
     #error := false;
     #status := #STATUS_FINISHED_NO_ERROR;
     #subfunctionStatus := #SUB_STATUS_NO_ERROR;
     // ENO mechanism is not used
     ENO := TRUE;
   END_REGION
END_FUNCTION

FUNCTION "LGF_RandomRange_Real" : Real   // FC10014, SCL
TITLE = LGF_RandomRange_Real
{ S7_Optimized_Access := 'TRUE' }
AUTHOR : Siemens_Digital_Industries
FAMILY : LGF
NAME : LGF_RandomRange_Real
// This function generates random numbers in defined limits (Datatype Real)
   VAR_INPUT
      minValue : Real;   // minimal Value random can reach / Minimum value of the range of the random number
      maxValue : Real;   // maximal Value random can reach / Maximum value of the range of the random number
   END_VAR
   VAR_OUTPUT
      error : Bool;   // Error if true
      status : Word;   // Status of the function
      subfunctionStatus : Word;   // Status or return value of called FB's, FCs and system blocks
   END_VAR
   VAR_TEMP
      tempTime : DTL;   // System time
      tempNanoSecondInDWord : DWord;   // UDINT converted to DWORD for access to individual bytes
      tempTimeStatus : Word;   // Status of the instruction RD_SYS_T
      tempRandomValue : DWord;   // Random-start-value
      tempNormReal : Real;   // normalized value
   END_VAR
   // Ret_Val : Returns random Real number in predefined range
   VAR CONSTANT
      ZERO : Real := 0.0;   // Zero value in case of error
      MAX_UDINT : UDInt := 4294967295;   // Maximum UDINT value
      SUB_STATUS_NO_ERROR : Word := 16#0000;   // Status: sub function call ends without error
      STATUS_FINISHED_NO_ERROR : Word := 16#0000;   // Status: Execution finished without errors
      ERR_MAX_LESS_MIN : Word := 16#8200;   // Error: The maximum limit number is smaller than the minimum limit number
      ERR_RD_SYS_T : Word := 16#8600;   // Error: System function Read system time returned an error
   END_VAR
BEGIN
   REGION Block info header
     //=============================================================================
     // SIEMENS AG / (c)Copyright 2017
     //-----------------------------------------------------------------------------
     // Title:            LGF_RandomRange_Real
     // Comment/Function: This function generates random numbers in defined limits (Datatype Real)
     // Library/Family:   LGF(Library General Functions)
     // Author:           Siemens Digital Industry Support
     // Tested with:      S7-PLCSIM Advanced V2.0 SP1
     // Engineering:      TIA Portal V15 Update 2
     // Restrictions:     ENO disabled - error handling done by error and status
     // Requirements:     PLC (S7-1200 / S7-1500)
     //-------------------------------------------------------------------------------
     // Change log table:
     // Version  | Date       | Expert in charge       | Changes applied
     //----------|------------|------------------------|------------------------------
     // 01.00.00 19.08.2015  Siemens Industry Online Support
     //                      First released version
     // 01.00.01 02.01.2017  Siemens Industry Online Support
     //                      Upgrade: TIA Portal V14 Update 1
     // 01.00.02 02.03.2017  Siemens Industry Online Support
     //                      Bugfix: FC number
     // 01.00.03 17.08.2018  Siemens Industry Online Support
     //                      Upgrade: TIA V15 Update 2
     // 01.00.04 23.11.2018  Siemens Industry Online Support
     //                      Upgrade: TIA V15.1
     // 01.01.00 13.11.2019  Siemens Industry Presales Support
     //                      Renamed from "LGF_RandomReal" to "LGF_RandomRange_Real"
     //                      Regions, commens and costants are added
     // 03.00.00 23.04.2020  Siemens Industry Support
     //                      Set version to V3.0.0, harmonize the version of the whole library
     //=============================================================================
   END_REGION

   REGION Validation
     // Check if the maximal Value is less than the minimal value
     IF (#minValue > #maxValue) THEN
       #error := true;
       #status := #ERR_MAX_LESS_MIN;
       #subfunctionStatus := #SUB_STATUS_NO_ERROR;
       #LGF_RandomRange_Real := #ZERO;
       RETURN;
     END_IF;

     // Read system time
     #tempTimeStatus := INT_TO_WORD(RD_SYS_T(#tempTime));

     // Check return variable for error
     IF (#tempTimeStatus <> #SUB_STATUS_NO_ERROR) THEN
       #error := true;
       #status := #ERR_RD_SYS_T;
       #subfunctionStatus := #tempTimeStatus;
       #LGF_RandomRange_Real := #ZERO;
       RETURN;
     END_IF;
   END_REGION

   REGION Calculating random number
     // Converting to double word so individual bytes can be addressed
     #tempNanoSecondInDWord := UDINT_TO_DWORD(#tempTime.NANOSECOND);

     // Calculate a random-start-value depending on the time
     #tempRandomValue.%B3 := #tempNanoSecondInDWord.%B0;
     #tempRandomValue.%B2 := #tempNanoSecondInDWord.%B1;
     #tempRandomValue.%B1 := #tempNanoSecondInDWord.%B2;
     #tempRandomValue.%B0 := #tempNanoSecondInDWord.%B3;

     // Norm the calculated random number: 0.0 <= #tempNormReal <= 1.0
     #tempNormReal := UDINT_TO_REAL(DWORD_TO_UDINT(#tempRandomValue)) / UDINT_TO_REAL(#MAX_UDINT);

     // Scale the tempNormReal to be in the range of maxValue and minValue
     #LGF_RandomRange_Real := ((#tempNormReal * (#maxValue - #minValue) + (#minValue)));

     #error := false;
     #status := #STATUS_FINISHED_NO_ERROR;
     #subfunctionStatus := #SUB_STATUS_NO_ERROR;
     // ENO mechanism is not used
     ENO := TRUE;
   END_REGION
END_FUNCTION

// folder: Library_LGF/6 Converter operations

FUNCTION "LGF_DTLtoString_ISO" : String   // FC10083, SCL
TITLE = LGF_DTLtoString_ISO
{ S7_Optimized_Access := 'TRUE' }
AUTHOR : Siemens_Industry_Online_Support
FAMILY : LGF
NAME : LGF_DTLtoString_ISO
// This function converts DTL into a string in ISO format.
   VAR_INPUT
      "date" : DTL;   // Date as DTL tag
      separator : Char;   // Separator between date components
   END_VAR
   VAR_TEMP
      tempString : String;   // temp string to setup the date string / -
      tempIndex : DInt;   // iterator for replacing withspaces with '0' in nanosecondstring / -
   END_VAR
   // Ret_Val : Date as String tag
   VAR CONSTANT
      CONVERT_SIZE_YEAR : USInt := 4;   // Number of character positions for Year
      CONVERT_SIZE_MONTH_DAY_HOUR_MINUTE_SECOND : USInt := 2;   // Number of character positions for Month, Day, Minute and Second
      CONVERT_SIZE_NANOSECOND : USInt := 9;   // Number of character positions for Nanoseconds
      CONVERT_PRECISION : USInt := 0;   // Number of decimal places to convert
      CONVERT_FORMAT_TO_STRING : Word := 16#0000;   // Output format of the characters
      CONVERT_START_POSITION_YEAR : UInt := 1;   // Character starting in string at which position the result is written.
      CONVERT_START_POSITION_MONTH : UInt := 6;   // Character starting in string at which position the result is written.
      CONVERT_START_POSITION_DAY : UInt := 9;   // Character starting in string at which position the result is written.
      CONVERT_START_POSITION_HOUR : UInt := 12;   // Character starting in string at which position the result is written.
      CONVERT_START_POSITION_MINUTE : UInt := 15;   // Character starting in string at which position the result is written.
      CONVERT_START_POSITION_SECOND : UInt := 18;   // Character starting in string at which position the result is written.
      CONVERT_START_POSITION_NANOSECOND : UInt := 21;   // Character starting in string at which position the result is written.
      SEPARATOR_POSITION_YEAR_MONTH : UInt := 5;   // Character starting in string at which position the result is written.
      SEPARATOR_POSITION_MONTH_DAY : UInt := 8;   // Character starting in string at which position the result is written.
      SEPARATOR_POSITION_HOUR_MINUTE : UInt := 14;   // Character starting in string at which position the result is written.
      SEPARATOR_POSITION_MINUTE_SECOND : UInt := 17;   // Character starting in string at which position the result is written.
      SEPARATOR_POSITION_SECOND_NANOSECOND : UInt := 20;   // Character starting in string at which position the result is written.
      SEPARATOR_NANOSECOND : Char := '.';   // Seperator for Nanosecond
      SEPARATOR_TIME : Char := ':';   // Seperator for Time
      SEPARATOR_DATE : Char := '-';   // Default separator for Date
      REPLACE_NANOSECOND_COUNT : DInt := 8;   // Number of Nonosecond characters to be checked for replacing withspaces wit '0'
   END_VAR
BEGIN
   REGION BLOCK INFO HEADER
     //===============================================================================
     // SIEMENS AG / (c)Copyright 2019
     //-------------------------------------------------------------------------------
     // Title:            LGF_DTLtoString_ISO
     // Comment/Function: This function converts DTL into a string in ISO format.
     // Library/Family:   LGF (Library General Functions)
     // Author:           Siemens Digital Industry Support
     // Tested with:      S7-PLCSIM Advanced V2.0 SP1
     // Engineering:      TIA Portal V15.1
     // Restrictions:     ENO mechanism is not used, no error handling
     // Requirements:     PLC (S7-1200 / S7-1500)
     //-------------------------------------------------------------------------------
     // Change log table:
     // Version  | Date       | Expert in charge       | Changes applied
     //----------|------------|------------------------|------------------------------
     // 01.00.00 | 15.06.2016 | Siemens Industry Online Support
     //                         First released version
     // 01.00.01 | 02.01.2017 | Siemens Industry Online Support
     //                         Upgrade: TIA Portal V14 Update 1
     // 01.00.02 | 17.08.2018 | Siemens Industry Online Support
     //                         Upgrade: TIA V15 Update 2
     // 01.00.03 | 23.11.2018 | Siemens Industry Online Support
     //                         Upgrade: TIA V15.1
     // 01.00.04 | 17.07.2019 | Siemens Industry Presale Support
     //                         BUgfix - nanosecond precision and '0' filling
     // 01.00.05 | 18.07.2019 | Siemens Industry Presale Support
     //                         renamed from "LGF_DTLtoString" to "LGF_DTLtoString_ISO"
     //                         split into two blocks, removed "format" input
     // 03.00.00 | 23.04.2020 | Siemens Industry Support | Set version to V3.0.0
     //                         harmonize the version of the whole library
     //=============================================================================
   END_REGION

   REGION INITIALISATION
     #tempString := '';
   END_REGION

   REGION CONVERTER
     // Set format parameters for output string
     // International ISO 8601
     // DTL  | Y| Y| Y| Y| -| M| M| -| D| D|  | H| H| :| M| M| :| S| S| .|NS|NS|NS|NS|NS|NS|NS|NS|NS
     // -----|--|--|--|--|--|--|--|--|--|--|--|--|--|--|--|--|--|--|--|--|--|--|--|--|--|--|--|--|--
     // Pos  | 1| 2| 3| 4| 5| 6| 7| 8| 9|10|11|12|13|14|15|16|17|18|19|20|21|22|23|24|25|26|27|28|29

     // Convert "Value" into "String" and place at the right position
     VAL_STRG(FORMAT := #CONVERT_FORMAT_TO_STRING,
              IN     := #date.YEAR,
              P      := #CONVERT_START_POSITION_YEAR,
              PREC   := #CONVERT_PRECISION,
              SIZE   := #CONVERT_SIZE_YEAR,
              OUT    => #tempString);    // DTL YEAR --> String --> #tempPosYear

     VAL_STRG(FORMAT := #CONVERT_FORMAT_TO_STRING,
              IN     := #date.MONTH,
              P      := #CONVERT_START_POSITION_MONTH,
              PREC   := #CONVERT_PRECISION,
              SIZE   := #CONVERT_SIZE_MONTH_DAY_HOUR_MINUTE_SECOND,
              OUT    => #tempString);     // DTL MONTH --> String --> #tempPosMonth

     VAL_STRG(FORMAT := #CONVERT_FORMAT_TO_STRING,
              IN     := #date.DAY,
              P      := #CONVERT_START_POSITION_DAY,
              PREC   := #CONVERT_PRECISION,
              SIZE   := #CONVERT_SIZE_MONTH_DAY_HOUR_MINUTE_SECOND,
              OUT    => #tempString);     // DTL DAY --> String --> #tempPosDay

     VAL_STRG(FORMAT := #CONVERT_FORMAT_TO_STRING,
              IN     := #date.HOUR,
              P      := #CONVERT_START_POSITION_HOUR,
              PREC   := #CONVERT_PRECISION,
              SIZE   := #CONVERT_SIZE_MONTH_DAY_HOUR_MINUTE_SECOND,
              OUT    => #tempString);     // DTL HOUR --> String --> #tempPosHour

     VAL_STRG(FORMAT := #CONVERT_FORMAT_TO_STRING,
              IN     := #date.MINUTE,
              P      := #CONVERT_START_POSITION_MINUTE,
              PREC   := #CONVERT_PRECISION,
              SIZE   := #CONVERT_SIZE_MONTH_DAY_HOUR_MINUTE_SECOND,
              OUT    => #tempString);     // DTL MINUTE --> String --> #tempPosMinute

     VAL_STRG(FORMAT := #CONVERT_FORMAT_TO_STRING,
              IN     := #date.SECOND,
              P      := #CONVERT_START_POSITION_SECOND,
              PREC   := #CONVERT_PRECISION,
              SIZE   := #CONVERT_SIZE_MONTH_DAY_HOUR_MINUTE_SECOND,
              OUT    => #tempString);     // DTL SECOND --> String --> #tempPosSecond

     VAL_STRG(FORMAT := #CONVERT_FORMAT_TO_STRING,
              IN     := #date.NANOSECOND,
              P      := #CONVERT_START_POSITION_NANOSECOND,
              PREC   := #CONVERT_PRECISION,
              SIZE   := #CONVERT_SIZE_NANOSECOND,
              OUT    => #tempString);     // DTL NANOSECOND --> String --> #tempPosNanosecond

     // Place separators at the right position in the string
     IF #separator = '' THEN
       #tempString[#SEPARATOR_POSITION_YEAR_MONTH] := #SEPARATOR_DATE;
       #tempString[#SEPARATOR_POSITION_MONTH_DAY] := #SEPARATOR_DATE;
     ELSE
       #tempString[#SEPARATOR_POSITION_YEAR_MONTH] := #separator;
       #tempString[#SEPARATOR_POSITION_MONTH_DAY] := #separator;
     END_IF;
     #tempString[#SEPARATOR_POSITION_HOUR_MINUTE] := #SEPARATOR_TIME;
     #tempString[#SEPARATOR_POSITION_MINUTE_SECOND] := #SEPARATOR_TIME;
     #tempString[#SEPARATOR_POSITION_SECOND_NANOSECOND] := #SEPARATOR_NANOSECOND;

     // Correcting the string, due to the conversion of a leading "0" value into a "blank".
     // Replacing of "blank" by "0"
     IF (#tempString[#CONVERT_START_POSITION_MONTH] = ' ') THEN
       #tempString[#CONVERT_START_POSITION_MONTH] := '0';
     END_IF;

     IF (#tempString[#CONVERT_START_POSITION_DAY] = ' ') THEN
       #tempString[#CONVERT_START_POSITION_DAY] := '0';
     END_IF;

     IF (#tempString[#CONVERT_START_POSITION_HOUR] = ' ') THEN
       #tempString[#CONVERT_START_POSITION_HOUR] := '0';
     END_IF;

     IF (#tempString[#CONVERT_START_POSITION_MINUTE] = ' ') THEN
       #tempString[#CONVERT_START_POSITION_MINUTE] := '0';
     END_IF;

     IF (#tempString[#CONVERT_START_POSITION_SECOND] = ' ') THEN
       #tempString[#CONVERT_START_POSITION_SECOND] := '0';
     END_IF;

     FOR #tempIndex := 0 TO #REPLACE_NANOSECOND_COUNT DO
       IF (#tempString[UINT_TO_SINT(#CONVERT_START_POSITION_NANOSECOND) + #tempIndex] = ' ') THEN
         #tempString[UINT_TO_SINT(#CONVERT_START_POSITION_NANOSECOND) + #tempIndex] := '0';
       ELSE
         EXIT;
       END_IF;
     END_FOR;
   END_REGION

   REGION OUTPUTS
     #LGF_DTLtoString_ISO := #tempString;
     // no error handling needed
     ENO := TRUE;
   END_REGION
END_FUNCTION

// folder: TaskErrors

ORGANIZATION_BLOCK "Time error interrupt"   // OB80, LAD, TimeErrorInterrupt
{ S7_Optimized_Access := 'TRUE' }
VERSION : 0.1
   VAR_INPUT
      Fault_ID : Byte;   // Fault identifier
      Csg_OBnr : OB_Any;   // Number of OB causing the error
      Csg_Prio : UInt;   // Priority of OB causing the error
   END_VAR
BEGIN
END_ORGANIZATION_BLOCK

ORGANIZATION_BLOCK "Diagnostic error interrupt"   // OB82, LAD, DiagnosticErrorInterrupt
{ S7_Optimized_Access := 'TRUE' }
VERSION : 0.1
   VAR_INPUT
      IO_State : Word;   // IO state of the HW object
      LADDR : Hw_Any;   // Hardware identifier
      Channel : UInt;   // Channel number
      MultiError : Bool;   // =true if more than one error is present
   END_VAR
   VAR_TEMP
      RALM : Struct
         AINFO : "AINFO_";
         TINFO : "TINFO_";
         RETVAL : Int;
         ALLARMI_da_OB82 : Struct
            RALM : "PN_Alarm";
            LADDR : Hw_Any;
            evento_uscente : Bool;
         END_STRUCT;
      END_STRUCT;
      TMP_dId : DInt;
   END_VAR
BEGIN

REGION Network 1
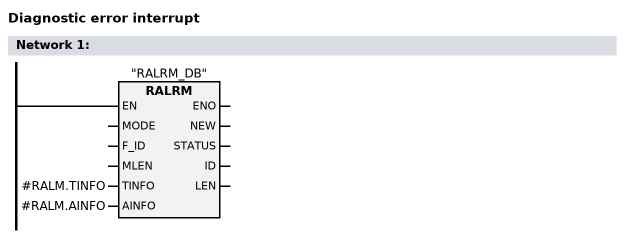
   "RALRM_DB"(TINFO := #RALM.TINFO, AINFO := #RALM.AINFO);   // RALRM
END_REGION

REGION Network 2 (SCL): Set alarms
   #TMP_dId:=UINT_TO_DINT("RALRM_DB".ID);

   IF "RALRM_DB".NEW THEN
       CASE #TMP_dId OF
           1:
               "RALRM_AUX_DB".tAlm.tF.xDevice1 := 1;
           2:
               "RALRM_AUX_DB".tAlm.tF.xDevice2 := 1;
           3:
               "RALRM_AUX_DB".tAlm.tF.xDevice3 := 1;
           4:
               "RALRM_AUX_DB".tAlm.tF.xDevice4 := 1;
           5:
               "RALRM_AUX_DB".tAlm.tF.xDevice5 := 1;
           6:
               "RALRM_AUX_DB".tAlm.tF.xDevice6 := 1;
           7:
               "RALRM_AUX_DB".tAlm.tF.xDevice7 := 1;
           8:
               "RALRM_AUX_DB".tAlm.tF.xDevice8 := 1;
           9:
               "RALRM_AUX_DB".tAlm.tF.xDevice9 := 1;
           10:
               "RALRM_AUX_DB".tAlm.tF.xDevice10 := 1;
           ELSE
               ;
       END_CASE;
   END_IF;
END_REGION
END_ORGANIZATION_BLOCK

ORGANIZATION_BLOCK "Pull or plug of modules"   // OB83, LAD, PullPlug
{ S7_Optimized_Access := 'TRUE' }
VERSION : 0.1
   VAR_INPUT
      LADDR : Hw_Io;   // Hardware identifier
      Event_Class : Byte;   // 16#38/39: module inserted, removed
      Fault_ID : Byte;   // Fault identifier
   END_VAR
BEGIN
END_ORGANIZATION_BLOCK

ORGANIZATION_BLOCK "Rack or station failure"   // OB86, LAD, RackStationFailure
{ S7_Optimized_Access := 'TRUE' }
VERSION : 0.1
   VAR_INPUT
      LADDR : Hw_Device;   // Hardware identifier
      Event_Class : Byte;   // Event class
      Fault_ID : Byte;   // Fault identifier
   END_VAR
BEGIN
END_ORGANIZATION_BLOCK

ORGANIZATION_BLOCK "Programming error"   // OB121, LAD, ProgrammingError
{ S7_Optimized_Access := 'TRUE' }
VERSION : 0.1
   VAR_INPUT
      BlockNr : UInt;   // Number of causing block
      Reaction : USInt;   // 0:ignore, 1:substitute, 2:skip
      Fault_ID : Byte;   // Fault identifier
      BlockType : USInt;   // 16#01:OB, 16#02:FC, 16#03:FB, 16#04:SFC, 16#05:SFB, 16#06:DB: Type of block causing the error
      Area : USInt;   // Area where the error occured
      DBNr : DB_ANY;   // DB number if Area = DB or DI
      Csg_OBNr : OB_Any;   // Number of OB causing the error
      Csg_Prio : USInt;   // Priority of OB causing the error
      Width : USInt;   // 0:bit, 1:byte, 2:word, 3:dword, 4:lword
   END_VAR
BEGIN
END_ORGANIZATION_BLOCK

ORGANIZATION_BLOCK "IO access error"   // OB122, LAD, IOAccessError
{ S7_Optimized_Access := 'TRUE' }
VERSION : 0.1
   VAR_INPUT
      BlockNr : UInt;   // Number of causing block
      Reaction : USInt;   // 0:ignore, 1:substitute, 2:skip
      Fault_ID : Byte;   // 16#42:reading, 16#43:writing
      BlockType : USInt;   // 16#01:OB, 16#02:FC, 16#03:FB, 16#04:SFC, 16#05:SFB, 16#06:DB: Type of block causing the error
      Area : USInt;   // 16#81:I, 16#82:Q: IO area where the IOaccess error occured
      DBNr : DB_ANY;   // Reserved for system
      Csg_OBNr : OB_Any;   // Number of OB causing the error
      Csg_Prio : USInt;   // Priority of OB causing the error
      Width : USInt;   // 0:bit, 1:byte, 2:word, 3:dword, 4:lword
   END_VAR
BEGIN
END_ORGANIZATION_BLOCK

// folder: TaskFast

ORGANIZATION_BLOCK "OBx_TaskFast"   // OB30, LAD, CyclicInterrupt
TITLE = Task fast OB
{ S7_Optimized_Access := 'TRUE' }
VERSION : 0.1
   VAR_INPUT
      Initial_Call : Bool;   // Initial call of this OB
      Event_Count : Int;   // Events discarded
   END_VAR
   VAR_TEMP
      TMP_lwDato : LWord;
      TMP_lrVal : LReal;
      TMP_rlVal : LReal;
      TMP_xValue : Bool;
      TMP_iRetVal : Int;
      TMP_stConnect : TCON_IP_v4;
   END_VAR
BEGIN

REGION Network 1: Initialize
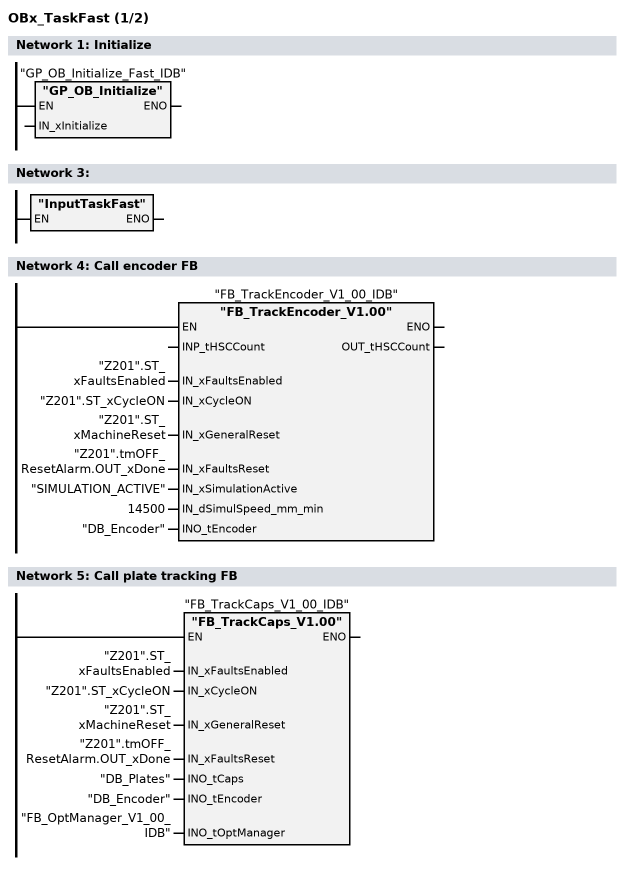
   RUNG wire#powerrail
      "GP_OB_Initialize_Fast_IDB"(IN_xInitialize :=)
   END_RUNG
   // the same network as SCL:
   "GP_OB_Initialize_Fast_IDB"();   // "GP_OB_Initialize"
END_REGION

REGION Network 2 (SCL): Message call

   "RP_OB_TaskFastToOpt"(FALSE);
   "RP_OB_TaskFastFromOpt"(FALSE);
END_REGION

REGION Network 3
   RUNG wire#powerrail
      "InputTaskFast"()
   END_RUNG
   // the same network as SCL:
   "InputTaskFast"();
END_REGION

REGION Network 4: Call encoder FB
   RUNG wire#powerrail
      "FB_TrackEncoder_V1_00_IDB"(INP_tHSCCount :=, IN_xFaultsEnabled := "Z201".ST_xFaultsEnabled, IN_xCycleON := "Z201".ST_xCycleON, IN_xGeneralReset := "Z201".ST_xMachineReset, IN_xFaultsReset := "Z201".tmOFF_ResetAlarm.OUT_xDone, IN_xSimulationActive := "SIMULATION_ACTIVE", IN_dSimulSpeed_mm_min := 14500, INO_tEncoder := "DB_Encoder", OUT_tHSCCount =>)
   END_RUNG
   // the same network as SCL:
   "FB_TrackEncoder_V1_00_IDB"(IN_xFaultsEnabled := "Z201".ST_xFaultsEnabled,   // "FB_TrackEncoder_V1.00"
                           IN_xCycleON := "Z201".ST_xCycleON,
                           IN_xGeneralReset := "Z201".ST_xMachineReset,
                           IN_xFaultsReset := "Z201".tmOFF_ResetAlarm.OUT_xDone,
                           IN_xSimulationActive := "SIMULATION_ACTIVE",
                           IN_dSimulSpeed_mm_min := 14500,
                           INO_tEncoder := "DB_Encoder");
END_REGION

REGION Network 5: Call plate tracking FB
   RUNG wire#powerrail
      "FB_TrackCaps_V1_00_IDB"(IN_xFaultsEnabled := "Z201".ST_xFaultsEnabled, IN_xCycleON := "Z201".ST_xCycleON, IN_xGeneralReset := "Z201".ST_xMachineReset, IN_xFaultsReset := "Z201".tmOFF_ResetAlarm.OUT_xDone, INO_tCaps := "DB_Plates", INO_tEncoder := "DB_Encoder", INO_tOptManager := "FB_OptManager_V1_00_IDB")
   END_RUNG
   // the same network as SCL:
   "FB_TrackCaps_V1_00_IDB"(IN_xFaultsEnabled := "Z201".ST_xFaultsEnabled,   // "FB_TrackCaps_V1.00"
                           IN_xCycleON := "Z201".ST_xCycleON,
                           IN_xGeneralReset := "Z201".ST_xMachineReset,
                           IN_xFaultsReset := "Z201".tmOFF_ResetAlarm.OUT_xDone,
                           INO_tCaps := "DB_Plates",
                           INO_tEncoder := "DB_Encoder",
                           INO_tOptManager := "FB_OptManager_V1_00_IDB");
END_REGION

REGION Network 6: Call defects tracking FB
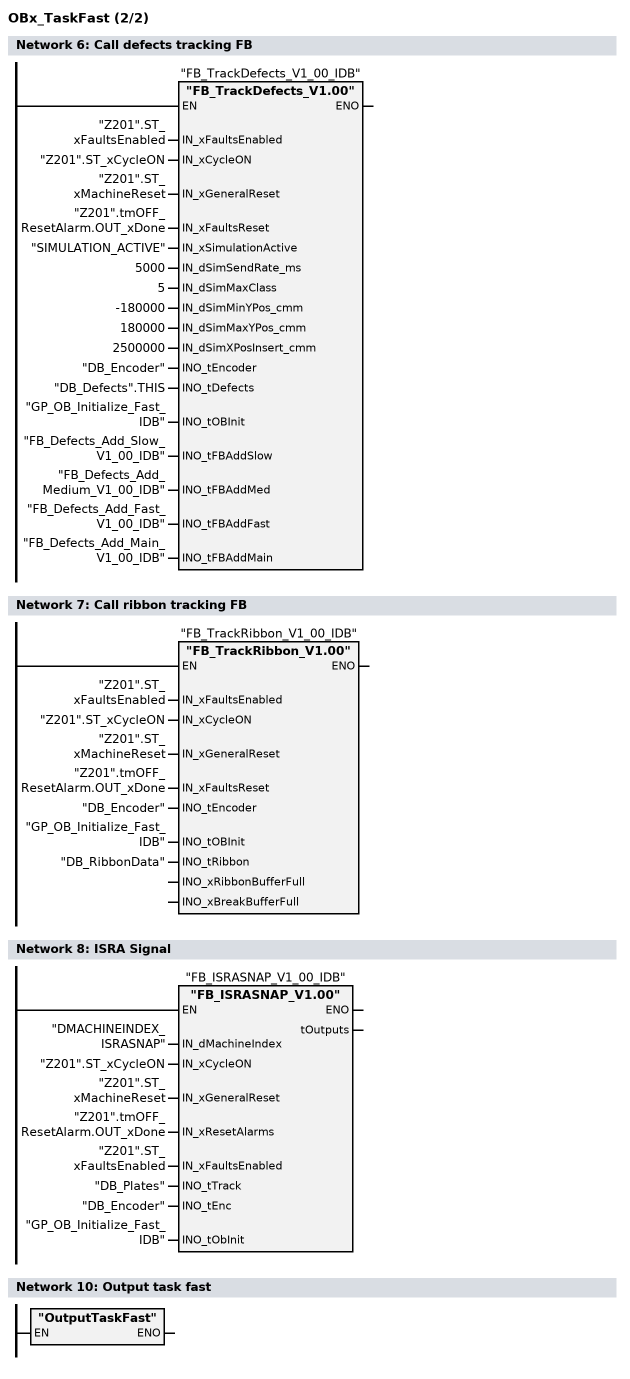
   RUNG wire#powerrail
      "FB_TrackDefects_V1_00_IDB"(IN_xFaultsEnabled := "Z201".ST_xFaultsEnabled, IN_xCycleON := "Z201".ST_xCycleON, IN_xGeneralReset := "Z201".ST_xMachineReset, IN_xFaultsReset := "Z201".tmOFF_ResetAlarm.OUT_xDone, IN_xSimulationActive := "SIMULATION_ACTIVE", IN_dSimSendRate_ms := 5000, IN_dSimMaxClass := 5, IN_dSimMinYPos_cmm := -180000, IN_dSimMaxYPos_cmm := 180000, IN_dSimXPosInsert_cmm := 2500000, INO_tEncoder := "DB_Encoder", INO_tDefects := "DB_Defects".THIS, INO_tOBInit := "GP_OB_Initialize_Fast_IDB", INO_tFBAddSlow := "FB_Defects_Add_Slow_V1_00_IDB", INO_tFBAddMed := "FB_Defects_Add_Medium_V1_00_IDB", INO_tFBAddFast := "FB_Defects_Add_Fast_V1_00_IDB", INO_tFBAddMain := "FB_Defects_Add_Main_V1_00_IDB")
   END_RUNG
   // the same network as SCL:
   "FB_TrackDefects_V1_00_IDB"(IN_xFaultsEnabled := "Z201".ST_xFaultsEnabled,   // "FB_TrackDefects_V1.00"
                           IN_xCycleON := "Z201".ST_xCycleON,
                           IN_xGeneralReset := "Z201".ST_xMachineReset,
                           IN_xFaultsReset := "Z201".tmOFF_ResetAlarm.OUT_xDone,
                           IN_xSimulationActive := "SIMULATION_ACTIVE",
                           IN_dSimSendRate_ms := 5000,
                           IN_dSimMaxClass := 5,
                           IN_dSimMinYPos_cmm := -180000,
                           IN_dSimMaxYPos_cmm := 180000,
                           IN_dSimXPosInsert_cmm := 2500000,
                           INO_tEncoder := "DB_Encoder",
                           INO_tDefects := "DB_Defects".THIS,
                           INO_tOBInit := "GP_OB_Initialize_Fast_IDB",
                           INO_tFBAddSlow := "FB_Defects_Add_Slow_V1_00_IDB",
                           INO_tFBAddMed := "FB_Defects_Add_Medium_V1_00_IDB",
                           INO_tFBAddFast := "FB_Defects_Add_Fast_V1_00_IDB",
                           INO_tFBAddMain := "FB_Defects_Add_Main_V1_00_IDB");
END_REGION

REGION Network 7: Call ribbon tracking FB
   RUNG wire#powerrail
      "FB_TrackRibbon_V1_00_IDB"(IN_xFaultsEnabled := "Z201".ST_xFaultsEnabled, IN_xCycleON := "Z201".ST_xCycleON, IN_xGeneralReset := "Z201".ST_xMachineReset, IN_xFaultsReset := "Z201".tmOFF_ResetAlarm.OUT_xDone, INO_tEncoder := "DB_Encoder", INO_tOBInit := "GP_OB_Initialize_Fast_IDB", INO_tRibbon := "DB_RibbonData", INO_xRibbonBufferFull :=, INO_xBreakBufferFull :=)
   END_RUNG
   // the same network as SCL:
   "FB_TrackRibbon_V1_00_IDB"(IN_xFaultsEnabled := "Z201".ST_xFaultsEnabled,   // "FB_TrackRibbon_V1.00"
                           IN_xCycleON := "Z201".ST_xCycleON,
                           IN_xGeneralReset := "Z201".ST_xMachineReset,
                           IN_xFaultsReset := "Z201".tmOFF_ResetAlarm.OUT_xDone,
                           INO_tEncoder := "DB_Encoder",
                           INO_tOBInit := "GP_OB_Initialize_Fast_IDB",
                           INO_tRibbon := "DB_RibbonData");
END_REGION

REGION Network 8: ISRA Signal
   RUNG wire#powerrail
      "FB_ISRASNAP_V1_00_IDB"(IN_dMachineIndex := "DMACHINEINDEX_ISRASNAP", IN_xCycleON := "Z201".ST_xCycleON, IN_xGeneralReset := "Z201".ST_xMachineReset, IN_xResetAlarms := "Z201".tmOFF_ResetAlarm.OUT_xDone, IN_xFaultsEnabled := "Z201".ST_xFaultsEnabled, INO_tTrack := "DB_Plates", INO_tEnc := "DB_Encoder", INO_tObInit := "GP_OB_Initialize_Fast_IDB", tOutputs =>)
   END_RUNG
   // the same network as SCL:
   "FB_ISRASNAP_V1_00_IDB"(IN_dMachineIndex := "DMACHINEINDEX_ISRASNAP",   // "FB_ISRASNAP_V1.00"
                           IN_xCycleON := "Z201".ST_xCycleON,
                           IN_xGeneralReset := "Z201".ST_xMachineReset,
                           IN_xResetAlarms := "Z201".tmOFF_ResetAlarm.OUT_xDone,
                           IN_xFaultsEnabled := "Z201".ST_xFaultsEnabled,
                           INO_tTrack := "DB_Plates",
                           INO_tEnc := "DB_Encoder",
                           INO_tObInit := "GP_OB_Initialize_Fast_IDB");
END_REGION

REGION Network 9 (SCL): Xcut
   #TMP_stConnect.ActiveEstablished := TRUE;
   #TMP_stConnect.ConnectionType := 11;    // TCP
   #TMP_stConnect.ID := "CONNUOC_XCUT1";
   #TMP_stConnect.InterfaceId := "Local~PROFINET_MCC1200";    // PROFINET Network
   #TMP_stConnect.LocalPort := 0;
   #TMP_stConnect.RemotePort := 502;   // 502 See TIA ONLINE HELP
   #TMP_stConnect.RemoteAddress.ADDR[1] := 192;
   #TMP_stConnect.RemoteAddress.ADDR[2] := 168;
   #TMP_stConnect.RemoteAddress.ADDR[3] := 21;
   #TMP_stConnect.RemoteAddress.ADDR[4] := 111;

   "FB_CrossCut1ModbusExchange_V1.00_DB"(IN_xGeneralReset := "Z201".ST_xMachineReset, IN_dMachineIndex := 0,
                                         INO_stConnect := #TMP_stConnect,
                                         INO_tMBClient := "DB_XCut1_MBClientInstance",
                                         INO_tXcut := "FB_CrossCuts_1_V1_00_IDB");

   #TMP_stConnect.ActiveEstablished := TRUE;
   #TMP_stConnect.ConnectionType := 11;    // TCP
   #TMP_stConnect.ID := "CONNUOC_XCUT2";
   #TMP_stConnect.InterfaceId := "Local~PROFINET_MCC1200";    // PROFINET Network
   #TMP_stConnect.LocalPort := 0;
   #TMP_stConnect.RemotePort := 502;   // 502 See TIA ONLINE HELP
   #TMP_stConnect.RemoteAddress.ADDR[1] := 192;
   #TMP_stConnect.RemoteAddress.ADDR[2] := 168;
   #TMP_stConnect.RemoteAddress.ADDR[3] := 21;
   #TMP_stConnect.RemoteAddress.ADDR[4] := 112;

   "FB_CrossCut2ModbusExchange_V1.00_DB"(IN_xGeneralReset := "Z201".ST_xMachineReset, IN_dMachineIndex := 1,
                                         INO_stConnect := #TMP_stConnect,
                                         INO_tMBClient := "DB_XCut2_MBClientInstance",
                                         INO_tXcut := "FB_CrossCuts_2_V1_00_IDB");


   #TMP_stConnect.ActiveEstablished := TRUE;
   #TMP_stConnect.ConnectionType := 11;    // TCP
   #TMP_stConnect.ID := "CONNUOC_XCUT3";
   #TMP_stConnect.InterfaceId := "Local~PROFINET_MCC1200";    // PROFINET Network
   #TMP_stConnect.LocalPort := 0;
   #TMP_stConnect.RemotePort := 502;   // 502 See TIA ONLINE HELP
   #TMP_stConnect.RemoteAddress.ADDR[1] := 192;
   #TMP_stConnect.RemoteAddress.ADDR[2] := 168;
   #TMP_stConnect.RemoteAddress.ADDR[3] := 21;
   #TMP_stConnect.RemoteAddress.ADDR[4] := 113;

   "FB_CrossCut3ModbusExchange_V1.00_DB"(IN_xGeneralReset := "Z201".ST_xMachineReset,
                                         IN_dMachineIndex := 1,
                                         INO_stConnect := #TMP_stConnect,
                                         INO_tMBClient := "DB_XCut3_MBClientInstance",
                                         INO_tXcut := "FB_CrossCuts_3_V1_00_IDB");
END_REGION

REGION Network 10: Output task fast
   RUNG wire#powerrail
      "OutputTaskFast"()
   END_RUNG
   // the same network as SCL:
   "OutputTaskFast"();
END_REGION
END_ORGANIZATION_BLOCK

// folder: TaskMain

ORGANIZATION_BLOCK "Main"   // OB1, LAD, ProgramCycle
TITLE = "Main Program Sweep (Cycle)"
{ S7_Optimized_Access := 'TRUE' }
VERSION : 0.1
   VAR_INPUT
      Initial_Call : Bool;   // Initial call of this OB
      Remanence : Bool;   // =True, if remanent data are available
   END_VAR
   VAR_TEMP
      tmp_xDummy : Bool;
      TMP_dIndex : DInt;
      TMP_iRetVal : Int;
      TMP_rgtMotorConfig : "UDT_MotorConfig";
   END_VAR
BEGIN

REGION Network 1: Initialize
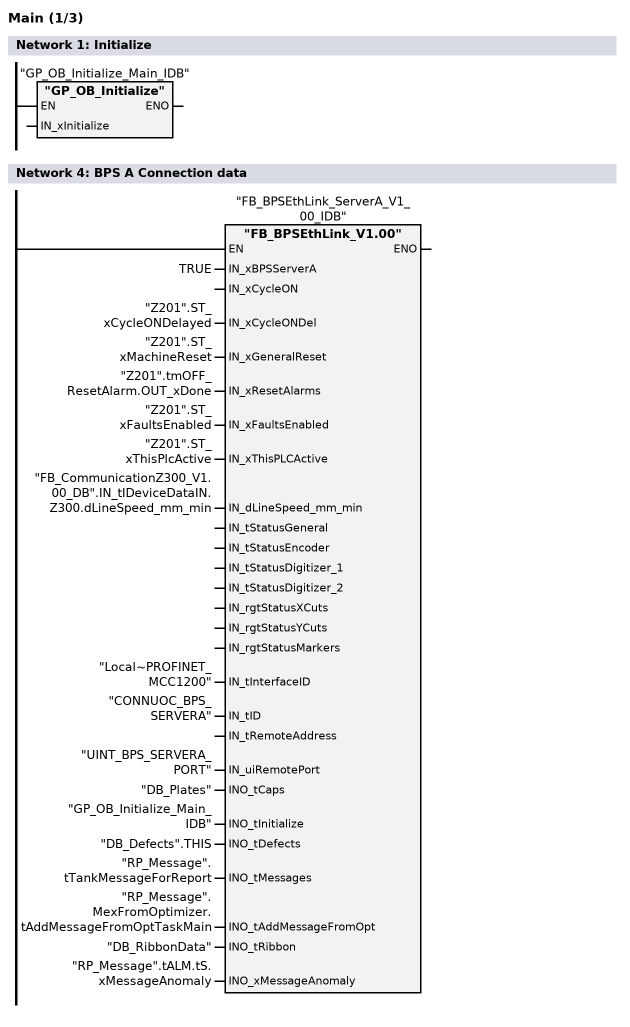
   RUNG wire#powerrail
      "GP_OB_Initialize_Main_IDB"(IN_xInitialize :=)
   END_RUNG
   // the same network as SCL:
   "GP_OB_Initialize_Main_IDB"();   // "GP_OB_Initialize"
END_REGION

REGION Network 2 (SCL): Message call

   "RP_OB_TaskMainToOpt"(FALSE);
   "RP_OB_TaskMainFromOpt"(FALSE);
END_REGION

REGION Network 3 (SCL): BPS Connection data ip
   //BPS Connection A

   "FB_BPSEthLink_ServerA_V1_00_IDB".IN_tRemoteAddress.ADDR[1] := "IPV4_BPS_SERVERA_IP1";
   "FB_BPSEthLink_ServerA_V1_00_IDB".IN_tRemoteAddress.ADDR[2] := "IPV4_BPS_SERVERA_IP2";
   "FB_BPSEthLink_ServerA_V1_00_IDB".IN_tRemoteAddress.ADDR[3] := "IPV4_BPS_SERVERA_IP3";
   "FB_BPSEthLink_ServerA_V1_00_IDB".IN_tRemoteAddress.ADDR[4] := "IPV4_BPS_SERVERA_IP4";

   "FB_BPSEthLink_ServerA_V1_00_IDB".IN_tStatusEncoder.dActualBTC_cmm := "DB_Encoder".dActualEncoderCounter_cmm;
   "FB_BPSEthLink_ServerA_V1_00_IDB".IN_tStatusEncoder.dTrackSpeed_mm_min := "DB_Encoder".dActSpeedValue_mm_min;